        [6]   // Conveyor 6 Millisecond Accumulator Updated by STI File 18
        [7]   // Conveyor 7 Millisecond Accumulator Updated by STI File 18
        [8]   // Conveyor 8 Millisecond Accumulator Updated by STI File 18
        [9]   // Conveyor 9 Millisecond Accumulator Updated by STI File 18
        [16]   // Conveyor 16 Millisecond Accumulator Updated by STI File 18
        [17]   // Conveyor 17 Millisecond Accumulator Updated by STI File 18
        [18]   // Conveyor 18 Millisecond Accumulator Updated by STI File 18
        [19]   // Conveyor 19 Millisecond Accumulator Updated by STI File 18
        [20]   // conveyor 20 Millisecond Accumulator Updated by STI File 18
        [21]   // conveyor 21 Millisecond Accumulator Updated by STI File 18
        [22]   // conveyor 22 Millisecond Accumulator Updated by STI File 18
        [23]   // conveyor 23 Millisecond Accumulator Updated by STI File 18
        [24]   // conveyor 24 Millisecond Accumulator Updated by STI File 18
        [25]   // conveyor 25 Millisecond Accumulator Updated by STI File 18
        [26]   // conveyor 26 Millisecond Accumulator Updated by STI File 18
        [27]   // conveyor 27 Millisecond Accumulator Updated by STI File 18
        [28]   // conveyor 28 Millisecond Accumulator Updated by STI File 18
        [29]   // conveyor 29 Millisecond Accumulator Updated by STI File 18
        [30]   // conveyor 30 Millisecond Accumulator Updated by STI File 18
        [31]   // conveyor 31 Millisecond Accumulator Updated by STI File 18
   N301 : DINT[1];
   N302 : DINT[1];
   N303 : DINT[1];
   N304 : DINT[1];
   N305 : DINT[1];
   N306 : DINT[1];
   N307 : DINT[1];
   N308 : DINT[1];
   N309 : DINT[1];
   N31 : DINT[33];   // M2 to M4
        [1]   // Conveyor 1 Copy Buffer Transfers PLC IDs to Next Conveyor
        [2]   // Conveyor 2 Copy Buffer Transfers PLC IDs to Next Conveyor
        [3]   // Conveyor 3 Copy Buffer Transfers PLC IDs to Next Conveyor
        [4]   // Conveyor 4 Copy Buffer Transfers PLC IDs to Next Conveyor
        [5]   // Conveyor 5 Copy Buffer Transfers PLC IDs to Next Conveyor
        [6]   // Conveyor 6 Copy Buffer Transfers PLC IDs to Next Conveyor
        [7]   // Conveyor 7 Copy Buffer Transfers PLC IDs to Next Conveyor
        [8]   // Conveyor 8 Copy Buffer Transfers PLC IDs to Next Conveyor
        [9]   // Conveyor 9 Copy Buffer Transfers PLC IDs to Next Conveyor
        [10]   // Conveyor 10 Copy Buffer Transfers PLC IDs to Next Conveyor
        [11]   // Conveyor 11 Copy Buffer Transfers PLC IDs to Next Conveyor
        [12]   // Conveyor 12 Copy Buffer Transfers PLC IDs to Next Conveyor
        [13]   // Conveyor 13 Copy Buffer Transfers PLC IDs to Next Conveyor
        [14]   // Conveyor 14 Copy Buffer Transfers PLC IDs to Next Conveyor
        [15]   // Conveyor 15 Copy Buffer Transfers PLC IDs to Next Conveyor
        [16]   // Conveyor 16 Copy Buffer Transfers PLC IDs to Next Conveyor
        [17]   // Conveyor 17 Copy Buffer Transfers PLC IDs to Next Conveyor
        [18]   // Conveyor 18 Copy Buffer Transfers PLC IDs to Next Conveyor
        [19]   // Conveyor 19 Copy Buffer Transfers PLC IDs to Next Conveyor
        [20]   // Conveyor 20 Copy Buffer Transfers PLC IDs to Next Conveyor
        [21]   // Conveyor 21 Copy Buffer Transfers PLC IDs to Next Conveyor
        [22]   // Conveyor 22 Copy Buffer Transfers PLC IDs to Next Conveyor
        [23]   // Conveyor 23 Copy Buffer Transfers PLC IDs to Next Conveyor
        [24]   // Conveyor 24 Copy Buffer Transfers PLC IDs to Next Conveyor
        [25]   // Conveyor 25 Copy Buffer Transfers PLC IDs to Next Conveyor
        [26]   // Conveyor 26 Copy Buffer Transfers PLC IDs to Next Conveyor
        [27]   // Conveyor 27 Copy Buffer Transfers PLC IDs to Next Conveyor
        [28]   // Conveyor 28 Copy Buffer Transfers PLC IDs to Next Conveyor
        [29]   // Conveyor 29 Copy Buffer Transfers PLC IDs to Next Conveyor
        [30]   // Conveyor 30 Copy Buffer Transfers PLC IDs to Next Conveyor
        [31]   // Conveyor 31 Copy Buffer Transfers PLC IDs to Next Conveyor
        [32]   // Conveyor 32 Copy Buffer Transfers PLC IDs to Next Conveyor
   N310 : DINT[1];
   N311 : DINT[1];
   N312 : DINT[1];
   N313 : DINT[1];
   N314 : DINT[1];
   N315 : DINT[1];
   N316 : DINT[1];
   N317 : DINT[1];
   N318 : DINT[1];
   N319 : DINT[1];
   N32 : DINT[33] := ([0] := 1800, [1] := 67);
        [10]   // Conveyor 10 Tracking Zone Length
        [11]   // Conveyor 11 Tracking Zone Length
        [12]   // Conveyor 12 Tracking Zone Length
        [13]   // Conveyor 13 Tracking Zone Length
        [1]   // Conveyor 1 Tracking Zone Length
        [14]   // Conveyor 14 Tracking Zone Length
        [2]   // Conveyor 2 Tracking Zone Length
        [15]   // Conveyor 15 Tracking Zone Length
        [3]   // Conveyor 3 Tracking Zone Length
        [16]   // Conveyor 16 Tracking Zone Length
        [17]   // Conveyor 17 Tracking Zone Length
        [18]   // Conveyor 18 Tracking Zone Length
        [19]   // Conveyor 19 Tracking Zone Length
        [20]   // Conveyor 20 Tracking Zone Length
        [21]   // Conveyor 21 Tracking Zone Length
        [22]   // Conveyor 22 Tracking Zone Length
        [23]   // Conveyor 23 Tracking Zone Length
        [24]   // Conveyor 24 Tracking Zone Length
        [25]   // Conveyor 25 Tracking Zone Length
        [26]   // Conveyor 26 Tracking Zone Length
        [4]   // Conveyor 4 Tracking Zone Length
        [27]   // Conveyor 27 Tracking Zone Length
        [28]   // Conveyor 28 Tracking Zone Length
        [29]   // Conveyor 29 Tracking Zone Length
        [30]   // Conveyor 30 Tracking Zone Length
        [31]   // Conveyor 31 Tracking Zone Length
        [32]   // Conveyor 32 Tracking Zone Length
        [5]   // Conveyor 5 Tracking Zone Length
        [6]   // Conveyor 6 Tracking Zone Length
        [7]   // Conveyor 7 Tracking Zone Length
        [8]   // Conveyor 8 Tracking Zone Length
        [9]   // Conveyor 9 Tracking Zone Length
   N320 : DINT[1];
   N321 : DINT[1];
   N322 : DINT[1];
   N323 : DINT[1];
   N324 : DINT[1];
   N325 : DINT[1];
   N326 : DINT[1];
   N327 : DINT[1];
   N328 : DINT[1];
   N329 : DINT[1];
   N33 : DINT[2] := ([0] := 3000, [1] := 40);
   N330 : DINT[1];
   N331 : DINT[1];
   N332 : DINT[1];
   N334 : DINT[1];
   N335 : DINT[1];
   N336 : DINT[1];
   N337 : DINT[1];
   N338 : DINT[1];
   N339 : DINT[1];
   N340 : DINT[1];
   N341 : DINT[1];
   N342 : DINT[1];
   N343 : DINT[1];
   N344 : DINT[1];
   N345 : DINT[1];
   N346 : DINT[1];
   N347 : DINT[1];
   N348 : DINT[1];
   N349 : DINT[1];
   N35 : DINT[5] := ([0] := 32, [1] := 232, [2] := 33, [3] := 132, [4] := 24);
   N350 : DINT[1];
   N351 : DINT[1];
   N352 : DINT[1];
   N353 : DINT[1];
   N354 : DINT[1];
   N355 : DINT[1];
   N356 : DINT[1];
   N357 : DINT[1];
   N358 : DINT[1];
   N359 : DINT[1];
   N35_0 : ALIAS FOR N35[0];
   N35_1 : ALIAS FOR N35[1];
   N35_2 : ALIAS FOR N35[2];
   N35_4 : ALIAS FOR N35[4];
   N360 : DINT[1];
   N361 : DINT[1];
   N362 : DINT[1];
   N363 : DINT[1];
   N364 : DINT[1];
   N365 : DINT[1];
   N367 : DINT[1];
   N368 : DINT[1];
   N369 : DINT[1];
   N370 : DINT[1];
   N371 : DINT[1];
   N372 : DINT[1];
   N373 : DINT[1];
   N374 : DINT[1];
   N375 : DINT[1];
   N376 : DINT[1];
   N377 : DINT[1];
   N378 : DINT[1];
   N379 : DINT[1];
   N380 : DINT[1];
   N381 : DINT[1];
   N382 : DINT[1];
   N383 : DINT[1];
   N384 : DINT[1];
   N385 : DINT[1];
   N386 : DINT[1];
   N387 : DINT[1];
   N388 : DINT[1];
   N389 : DINT[1];
   N390 : DINT[1];
   N391 : DINT[1];
   N392 : DINT[1];
   N393 : DINT[1];
   N394 : DINT[1];
   N395 : DINT[1];
   N396 : DINT[1];
   N397 : DINT[1];
   N398 : DINT[1];
   N40 : DINT[32];
        [10]   // Conveyor 10 PLD ID of Cap being Resynced
        [11]   // Conveyor 11 PLD ID of Cap being Resynced
        [12]   // Conveyor 12 PLD ID of Cap being Resynced
        [13]   // Conveyor 13 PLD ID of Cap being Resynced
        [14]   // Conveyor 14 PLD ID of Cap being Resynced
        [15]   // Conveyor 15 PLD ID of Cap being Resynced
        [16]   // Conveyor 16 PLD ID of Cap being Resynced
        [17]   // Conveyor 17 PLD ID of Cap being Resynced
        [18]   // Conveyor 18 PLD ID of Cap being Resynced
        [19]   // Conveyor 19 PLD ID of Cap being Resynced
        [20]   // Conveyor 20 PLD ID of Cap being Resynced
        [21]   // Conveyor 21 PLD ID of Cap being Resynced
        [22]   // Conveyor 22 PLD ID of Cap being Resynced
        [23]   // Conveyor 23 PLD ID of Cap being Resynced
        [24]   // Conveyor 24 PLD ID of Cap being Resynced
        [25]   // Conveyor 25 PLD ID of Cap being Resynced
        [26]   // Conveyor 26 PLD ID of Cap being Resynced
        [27]   // Conveyor 27 PLD ID of Cap being Resynced
        [28]   // Conveyor 28 PLD ID of Cap being Resynced
        [29]   // Conveyor 29 PLD ID of Cap being Resynced
        [1]   // Conveyor 1 PLD ID of Cap being Resynced
        [2]   // Conveyor 2 PLD ID of Cap being Resynced
        [3]   // Conveyor 3 PLD ID of Cap being Resynced
        [4]   // Conveyor 4 PLD ID of Cap being Resynced
        [5]   // Conveyor 5 PLD ID of Cap being Resynced
        [6]   // Conveyor 6 PLD ID of Cap being Resynced
        [7]   // Conveyor 7 PLD ID of Cap being Resynced
        [8]   // Conveyor 8 PLD ID of Cap being Resynced
        [9]   // Conveyor 9 PLD ID of Cap being Resynced
        [30]   // Conveyor 30 PLD ID of Cap being Resynced
        [31]   // Conveyor 31 PLD ID of Cap being Resynced
   N400 : DINT[1];
   N401 : DINT[1];
   N402 : DINT[1];
   N403 : DINT[1];
   N404 : DINT[1];
   N405 : DINT[1];
   N406 : DINT[1];
   N407 : DINT[1];
   N408 : DINT[1];
   N409 : DINT[1];
   N410 : DINT[1];
   N411 : DINT[1];
   N412 : DINT[1];
   N413 : DINT[1];
   N414 : DINT[1];
   N415 : DINT[1];
   N416 : DINT[1];
   N417 : DINT[1];
   N418 : DINT[1];
   N419 : DINT[1];
   N420 : DINT[1];
   N421 : DINT[1];
   N422 : DINT[1];
   N423 : DINT[1];
   N424 : DINT[1];
   N425 : DINT[1];
   N426 : DINT[1];
   N427 : DINT[1];
   N428 : DINT[1];
   N429 : DINT[1];
   N430 : DINT[1];
   N431 : DINT[1];
   N433 : DINT[1];
   N434 : DINT[1];
   N435 : DINT[1];
   N436 : DINT[1];
   N437 : DINT[1];
   N438 : DINT[1];
   N439 : DINT[1];
   N440 : DINT[1];
   N441 : DINT[1];
   N442 : DINT[1];
   N443 : DINT[1];
   N444 : DINT[1];
   N445 : DINT[1];
   N446 : DINT[1];
   N447 : DINT[1];
   N448 : DINT[1];
   N449 : DINT[1];
   N450 : DINT[1];
   N451 : DINT[1];
   N452 : DINT[1];
   N453 : DINT[1];
   N454 : DINT[1];
   N455 : DINT[1];
   N456 : DINT[1];
   N457 : DINT[1];
   N458 : DINT[1];
   N459 : DINT[1];
   N460 : DINT[1];
   N461 : DINT[1];
   N462 : DINT[1];
   N463 : DINT[1];
   N464 : DINT[1];
   N466 : DINT[1];
   N467 : DINT[1];
   N468 : DINT[1];
   N469 : DINT[1];
   N470 : DINT[1];
   N471 : DINT[1];
   N472 : DINT[1];
   N473 : DINT[1];
   N474 : DINT[1];
   N475 : DINT[1];
   N476 : DINT[1];
   N477 : DINT[1];
   N478 : DINT[1];
   N479 : DINT[1];
   N480 : DINT[1];
   N481 : DINT[1];
   N482 : DINT[1];
   N483 : DINT[1];
   N484 : DINT[1];
   N485 : DINT[1];
   N486 : DINT[1];
   N487 : DINT[1];
   N488 : DINT[1];
   N489 : DINT[1];
   N490 : DINT[1];
   N491 : DINT[1];
   N492 : DINT[1];
   N493 : DINT[1];
   N494 : DINT[1];
   N495 : DINT[1];
   N496 : DINT[1];
   N497 : DINT[1];
   N500 : DINT[13] := ([1] := 1755, [2] := 1755, [3] := 1750, [4] := 1750, [5] := 1750, [6] := 1750, [7] := 1750, [8] := 1755, [9] := 1755, [10] := 1755, [11] := 1755, [12] := 1755);   // Motor RPM
        [10]   // M2CM10 Motor RPM
        [11]   // M2CM11 Motor RPM
        [12]   // M2CM12 Motor RPM
        [1]   // M2CM01 Motor RPM
        [2]   // M2CM02 Motor RPM
        [3]   // M2CM03 Motor RPM
        [4]   // M2CM04 Motor RPM
        [5]   // M2CM05 Motor RPM
        [6]   // M2CM06 Motor RPM
        [7]   // M2CM07 Motor RPM
        [8]   // M2CM08 Motor RPM
        [9]   // M2CM09 Motor RPM
   N501 : DINT[13] := ([1] := 43, [2] := 43, [3] := 43, [4] := 29, [5] := 29, [6] := 29, [7] := 29, [8] := 29, [9] := 29, [10] := 29, [11] := 29, [12] := 29);   // Gearbox raito
        [10]   // M2CM10 Gearbox raito
        [11]   // M2CM11 Gearbox raito
        [12]   // M2CM12 Gearbox raito
        [1]   // M2CM01 Gearbox raito
        [2]   // M2CM02 Gearbox raito
        [3]   // M2CM03 Gearbox raito
        [4]   // M2CM04 Gearbox raito
        [5]   // M2CM05 Gearbox raito
        [6]   // M2CM06 Gearbox raito
        [7]   // M2CM07 Gearbox raito
        [8]   // M2CM08 Gearbox raito
        [9]   // M2CM09 Gearbox raito
   N502 : DINT[13] := ([1] := 100, [2] := 100, [3] := 100, [4] := 100, [5] := 100, [6] := 100, [7] := 100, [8] := 100, [9] := 100, [10] := 100, [11] := 100, [12] := 100);   // Slip compensation
        [10]   // M2 CM10 Slip Compensation
        [11]   // M2 CM11 Slip Compensation
        [12]   // M2 CM12 Slip Compensation
        [1]   // M2 CM01 Slip Compensation
        [2]   // M2 CM02 Slip Compensation
        [3]   // M2 CM03 Slip Compensation
        [4]   // M2 CM04 Slip Compensation
        [5]   // M2 CM05 Slip Compensation
        [6]   // M2 CM06 Slip Compensation
        [7]   // M2 CM07 Slip Compensation
        [8]   // M2 CM08 Slip Compensation
        [9]   // M2 CM09 Slip Compensation
   N504 : DINT[13] := ([1] := 2042, [2] := 2042, [3] := 1728, [4] := 1728, [5] := 1728, [6] := 1728, [7] := 1728, [8] := 1728, [9] := 1728, [10] := 1728, [11] := 1728, [12] := 1728);   // Roll Circ
        [10]   // M2CM10 Roll Circ
        [11]   // M2CM11 Roll Circ
        [12]   // M2CM12 Roll Circ
        [1]   // M2CM01 Roll Circ
        [2]   // M2CM02 Roll Circ
        [3]   // M2CM03 Roll Circ
        [4]   // M2CM04 Roll Circ
        [5]   // M2CM05 Roll Circ
        [6]   // M2CM06 Roll Circ
        [7]   // M2CM07 Roll Circ
        [8]   // M2CM08 Roll Circ
        [9]   // M2CM09 Roll Circ
   N505 : DINT[13] := ([1] := 1397, [2] := 1397, [3] := 1179, [4] := 1748, [5] := 1748, [6] := 1748, [7] := 1748, [8] := 1753, [9] := 1753, [10] := 1753, [11] := 1753, [12] := 1753);   // IPM/HZ Conv Factor
        [10]   // M2CM10 IPM/HZ Conv Factor
        [11]   // M2CM11 IPM/HZ Conv Factor
        [12]   // M2CM12 IPM/HZ Conv Factor
        [1]   // M2CM01 IPM/HZ Conv Factor
        [2]   // M2CM02 IPM/HZ Conv Factor
        [3]   // M2CM03 IPM/HZ Conv Factor
        [4]   // M2CM04 IPM/HZ Conv Factor
        [5]   // M2CM05 IPM/HZ Conv Factor
        [6]   // M2CM06 IPM/HZ Conv Factor
        [7]   // M2CM07 IPM/HZ Conv Factor
        [8]   // M2CM08 IPM/HZ Conv Factor
        [9]   // M2CM09 IPM/HZ Conv Factor
   N507 : DINT[26] := ([1] := 94, [2] := 94, [3] := 112, [4] := 76, [5] := 76, [6] := 76, [7] := 76, [8] := 75, [9] := 75, [10] := 75, [11] := 75, [12] := 75, [13] := 322, [14] := 322, [15] := 382, [16] := 257, [17] := 257, [18] := 257, [19] := 257, [20] := 257, [21] := 257, [22] := 257, [23] := 257, [24] := 257, [25] := 450);   // Drive Command HZ
        [7]   // M2CM07S A1 Data In
   N54 : DINT[251];
   N601 : DINT[25];
   N602 : DINT[25];
   N603 : DINT[25];
   N604 : DINT[25];
   N605 : DINT[25];
   N606 : DINT[25];
   N607 : DINT[25];
   N608 : DINT[25];
   N609 : DINT[25];
   N610 : DINT[25];
   N611 : DINT[25];
   N612 : DINT[25];
   N613 : DINT[25];
   N614 : DINT[25];
   N615 : DINT[25];
   N616 : DINT[25];
   N617 : DINT[25];
   N618 : DINT[25];
   N619 : DINT[25];
   N620 : DINT[25];
   N621 : DINT[25];
   N622 : DINT[25];
   N623 : DINT[25];
   N624 : DINT[25];
   N625 : DINT[25];
   N626 : DINT[25];
   N627 : DINT[25];
   N628 : DINT[25];
   N629 : DINT[25];
   N630 : DINT[25];
   N631 : DINT[25];
   N632 : DINT[25];
   N633 : DINT[25];
   N634 : DINT[25];
   N635 : DINT[25];
   N636 : DINT[25];
   N637 : DINT[25];
   N638 : DINT[25];
   N639 : DINT[25];
   N640 : DINT[25];
   N641 : DINT[25];
   N642 : DINT[25];
   N643 : DINT[25];
   N644 : DINT[25];
   N645 : DINT[25];
   N646 : DINT[25];
   N647 : DINT[25];
   N648 : DINT[25];
   N649 : DINT[25];
   N650 : DINT[25];
   N651 : DINT[25];
   N652 : DINT[25];
   N653 : DINT[25];
   N654 : DINT[25];
   N655 : DINT[25];
   N656 : DINT[25];
   N657 : DINT[25];
   N658 : DINT[25];
   N659 : DINT[25];
   N660 : DINT[25];
   N662 : DINT[25];
   N663 : DINT[25];
   N664 : DINT[25];
   N665 : DINT[25];
   N666 : DINT[25];
   N667 : DINT[25];
   N668 : DINT[25];
   N669 : DINT[25];
   N670 : DINT[25];
   N671 : DINT[25];
   N672 : DINT[25];
   N673 : DINT[25];
   N674 : DINT[25];
   N675 : DINT[25];
   N676 : DINT[25];
   N677 : DINT[25];
   N678 : DINT[25];
   N679 : DINT[25];
   N680 : DINT[25];
   N681 : DINT[25];
   N682 : DINT[25];
   N683 : DINT[25];
   N684 : DINT[25];
   N685 : DINT[25];
   N686 : DINT[25];
   N687 : DINT[25];
   N688 : DINT[25];
   N689 : DINT[25];
   N690 : DINT[25];
   N691 : DINT[25];
   N692 : DINT[25];
   N693 : DINT[25];
   N694 : DINT[25];
   N695 : DINT[25];
   N696 : DINT[25];
   N697 : DINT[25];
   N698 : DINT[25];
   N699 : DINT[25];
   N7 : DINT[101] := ([10] := 3500, [11] := 100, [20] := 3930);
        [10]   // Current Command Frequency
        [0]   // DH+ Station number set on processor DIP switches
        [11]   // Current Test Addition Operand
   N70 : DINT[128] := ([0] := 11008);
   N700 : DINT[25];
   N701 : DINT[25];
   N702 : DINT[25];
   N703 : DINT[25];
   N704 : DINT[25];
   N705 : DINT[25];
   N706 : DINT[25];
   N707 : DINT[25];
   N708 : DINT[25];
   N709 : DINT[25];
   N71 : DINT[128] := ([2] := 40, [4] := 60);
        [2]   // M2CM12 A1 Data In
        [4]   // M2CM12 A2 Data In
   N710 : DINT[25];
   N711 : DINT[25];
   N712 : DINT[25];
   N713 : DINT[25];
   N714 : DINT[25];
   N715 : DINT[25];
   N716 : DINT[25];
   N717 : DINT[25];
   N718 : DINT[25];
   N719 : DINT[25];
   N72 : DINT[200] := ([0] := 4095);
        [0].0   // M2CM01 Drive Healthy and Running
        [0].1   // M2CM02 Drive Healthy and Running
        [0].2   // M2CM03 Drive Healthy and Running
        [3]   // VMCC M2 Drive Fault or Not Running Bits NORTH
        [0]   // VMCC M2 Drive Status Word Drive Healthy
        [1]   // VMCC M2 Drive Fault or Not Running Bits
        [0].10   // M2CM11 Drive Healthy and Running
        [0].11   // M2CM12 Drive Healthy and Running
        [2].10   // M2CM11N Drive Healthy and Running
        [2].11   // M2CM12N Drive Healthy and Running
        [0].3   // M2CM04 Drive Healthy and Running
        [0].4   // M2CM05 Drive Healthy and Running
        [0].5   // M2CM06 Drive Healthy and Running
        [0].6   // M2CM07 Drive Healthy and Running
        [0].7   // M2CM08 Drive Healthy and Running
        [0].8   // M2CM09 Drive Healthy and Running
        [0].9   // M2CM10 Drive Healthy and Running
        [2].3   // M2CM04N Drive Healthy and Running
        [2].4   // M2CM05N Drive Healthy and Running
        [2].5   // M2CM06N Drive Healthy and Running
        [2].6   // M2CM07N Drive Healthy and Running
        [2].7   // M2CM08N Drive Healthy and Running
        [2].8   // M2CM09N Drive Healthy and Running
        [2].9   // M2CM10N Drive Healthy and Running
   N720 : DINT[25];
   N721 : DINT[25];
   N723 : DINT[25];
   N724 : DINT[25];
   N725 : DINT[25];
   N726 : DINT[25];
   N727 : DINT[25];
   N728 : DINT[25];
   N729 : DINT[25];
   N730 : DINT[25];
   N731 : DINT[25];
   N732 : DINT[25];
   N733 : DINT[25];
   N734 : DINT[25];
   N735 : DINT[25];
   N736 : DINT[25];
   N737 : DINT[25];
   N738 : DINT[25];
   N739 : DINT[25];
   N740 : DINT[25];
   N741 : DINT[25];
   N742 : DINT[25];
   N743 : DINT[25];
   N744 : DINT[25];
   N745 : DINT[25];
   N746 : DINT[25];
   N747 : DINT[25];
   N748 : DINT[25];
   N749 : DINT[25];
   N750 : DINT[25];
   N751 : DINT[25];
   N752 : DINT[25];
   N753 : DINT[25];
   N754 : DINT[25];
   N755 : DINT[25];
   N756 : DINT[25];
   N758 : DINT[25];
   N759 : DINT[25];
   N760 : DINT[25];
   N761 : DINT[25];
   N762 : DINT[25];
   N763 : DINT[25];
   N764 : DINT[25];
   N765 : DINT[25];
   N766 : DINT[25];
   N767 : DINT[25];
   N768 : DINT[25];
   N769 : DINT[25];
   N770 : DINT[25];
   N771 : DINT[25];
   N772 : DINT[25];
   N773 : DINT[25];
   N774 : DINT[25];
   N775 : DINT[25];
   N776 : DINT[25];
   N777 : DINT[25];
   N778 : DINT[25];
   N779 : DINT[25];
   N780 : DINT[25];
   N781 : DINT[25];
   N782 : DINT[25];
   N783 : DINT[25];
   N784 : DINT[25];
   N785 : DINT[25];
   N786 : DINT[25];
   N787 : DINT[25];
   N788 : DINT[25];
   N789 : DINT[25];
   N790 : DINT[25];
   N791 : DINT[25];
   N792 : DINT[25];
   N793 : DINT[25];
   N794 : DINT[25];
   N795 : DINT[25];
   N796 : DINT[25];
   N797 : DINT[25];
   N798 : DINT[25];
   N799 : DINT[25];
   N80 : DINT[65] := ([11] := 2415, [12] := 5642, [15] := 2284, [16] := 5646, [19] := 1825, [20] := 4512, [23] := 1683, [24] := 4510, [27] := 1685, [28] := 4515, [31] := 1682, [32] := 4517, [35] := 1697, [36] := 452, [39] := 1681, [40] := 2811, [43] := 1681, [44] := 2811, [47] := 1681, [48] := 2811, [51] := 1684, [52] := 2815, [55] := 3995, [56] := 5974, [60] := 3000, [64] := 3000);
        [13].8   // M2CM02 Accel Time
        [1]   // RIO SN WRITE DATA Reserved Not Used
        [13].9   // M2CM02 Accel Time
        [2]   // RIO SN WRITE DATA Reserved Not Used
        [13].1   // M2CM02 Start
        [13]   // M2CM02 Drive Command
        [3]   // RIO SN WRITE DATA Reserved Not Used
        [4]   // RIO SN WRITE DATA Reserved Not Used
        [13].6   // M2CM02 Local
        [17].1   // M2CM03 Start
        [9].8   // M2CM01 Accel Time
        [9].9   // M2CM01 Accel Time
        [13].7   // M2CM02 MOP Increment
        [10]   // M2CM01 Speed Reference
        [5]   // RIO SN WRITE DATA Reserved Not Used
        [6]   // RIO SN WRITE DATA Reserved Not Used
        [7]   // RIO SN WRITE DATA Reserved Not Used
        [13].15   // M2CM02 MOP Decrement
        [8]   // RIO SN WRITE DATA Reserved Not Used
        [17].8   // M2CM03 Accel Time
        [17].15   // M2CM03 MOP Decrement
        [21].15   // M2CM04 MOP Decrement
        [25].15   // M2CM05 MOP Decrement
        [18].1   // M2CM03 Reference Select
        [13].12   // M2CM02 Reference Select
        [13].13   // M2CM02 Reference Select
        [13].14   // M2CM02 Reference Select
        [13].0   // M2CM02 Stop
        [17].0   // M2CM03 Stop
        [14]   // M2CM02 Speed Reference
        [11]   // M2CM01 A1 Data In
        [12]   // M2CM01 A2 Data In
        [13].4   // M2CM02 Direction
        [21].0   // M2CM04 Stop
        [17].6   // M2CM03 Local
        [13].10   // M2CM02 Decel Time
        [13].11   // M2CM02 Decel Time
        [17].12   // M2CM03 Reference Select
        [17].13   // M2CM03 Reference Select
        [17].14   // M2CM03 Reference Select
        [29].15   // M2CM06 MOP Decrement
        [13].2   // M2CM02 Jog
        [13].3   // M2CM02 Clear Faults
        [13].5   // M2CM02 Direction
        [17]   // M2CM03 Drive Command
        [21].1   // M2CM04 Start
        [17].7   // M2CM03 MOP Increment
        [17].9   // M2CM03 Accel Time
        [21].8   // M2CM04 Accel Time
        [18]   // M2CM03 Speed Reference
        [15]   // M2CM02 A1 Data In
        [16]   // M2CM02 A2 Data In
        [17].4   // M2CM03 Direction
        [25].0   // M2CM05 Stop
        [21].6   // M2CM04 Local
        [17].10   // M2CM03 Decel Time
        [17].11   // M2CM03 Decel Time
        [21].12   // M2CM04 Reference Select
        [21].13   // M2CM04 Reference Select
        [21].14   // M2CM04 Reference Select
        [33].15   // M2CM07 MOP Decrement
        [17].2   // M2CM03 Jog
        [17].3   // M2CM03 Clear Faults
        [17].5   // M2CM03 Direction
        [21]   // M2CM04 Drive Command
        [25].1   // M2CM05 Start
        [21].7   // M2CM04 MOP Increment
        [21].9   // M2CM04 Accel Time
        [25].8   // M2CM05 Accel Time
        [22]   // M2CM04 Speed Reference
        [22].5   // M2CM04 Reference Select
        [19]   // M2CM03 A1 Data In
        [20]   // M2CM03 A2 Data In
        [21].4   // M2CM04 Direction
        [29].0   // M2CM06 Stop
        [25].6   // M2CM05 Local
        [21].10   // M2CM04 Decel Time
        [21].11   // M2CM04 Decel Time
        [25].12   // M2CM05 Reference Select
        [25].13   // M2CM05 Reference Select
        [25].14   // M2CM05 Reference Select
        [37].15   // M2CM08 MOP Decrement
        [21].2   // M2CM04 Jog
        [21].3   // M2CM04 Clear Faults
        [21].5   // M2CM04 Direction
        [25]   // M2CM05 Drive Command
        [29].1   // M2CM06 Start
        [25].7   // M2CM05 MOP Increment
        [25].9   // M2CM05 Accel Time
        [29].8   // M2CM06 Accel Time
        [26]   // M2CM05 Speed Reference
        [26].9   // M2CM05 Reference Select
        [23]   // M2CM04 A1 Data In
        [24]   // M2CM04 A2 Data In
        [25].4   // M2CM05 Direction
        [33].0   // M2CM07 Stop
        [29].6   // M2CM06 Local
        [25].10   // M2CM05 Decel Time
        [25].11   // M2CM05 Decel Time
        [29].12   // M2CM06 Reference Select
        [29].13   // M2CM06 Reference Select
        [29].14   // M2CM06 Reference Select
        [41].15   // M2CM09 MOP Decrement
        [25].2   // M2CM05 Jog
        [25].3   // M2CM05 Clear Faults
        [25].5   // M2CM05 Direction
        [29]   // M2CM06 Drive Command
        [33].1   // M2CM07 Start
        [29].7   // M2CM06 MOP Increment
        [29].9   // M2CM06 Accel Time
        [33].8   // M2CM07 Accel Time
        [30]   // M2CM06 Speed Reference
        [35].1   // M2CM07 Reference Select
        [27]   // M2CM05 A1 Data In
        [28]   // M2CM05 A2 Data In
        [29].4   // M2CM06 Direction
        [37].0   // M2CM08 Stop
        [33].6   // M2CM07 Local
        [29].10   // M2CM06 Decel Time
        [29].11   // M2CM06 Decel Time
        [30].13   // M2CM06 Reference Select
        [33].12   // M2CM07 Reference Select
        [33].13   // M2CM07 Reference Select
        [45].15   // M2CM10 MOP Decrement
        [29].2   // M2CM06 Jog
        [29].3   // M2CM06 Clear Faults
        [29].5   // M2CM06 Direction
        [33]   // M2CM07 Drive Command
        [37].1   // M2CM08 Start
        [33].7   // M2CM07 MOP Increment
        [33].9   // M2CM07 Accel Time
        [37].8   // M2CM08 Accel Time
        [34]   // M2CM07 Speed Reference
        [33].14   // M2CM07 Reference Select
        [31]   // M2CM06 A1 Data In
        [32]   // M2CM06 A2 Data In
        [33].4   // M2CM07 Direction
        [41].0   // M2CM09 Stop
        [37].6   // M2CM08 Local
        [33].10   // M2CM07 Decel Time
        [33].11   // M2CM07 Decel Time
        [37].12   // M2CM08 Reference Select
        [37].13   // M2CM08 Reference Select
        [37].14   // M2CM08 Reference Select
        [49].15   // M2CM11 MOP Decrement
        [33].2   // M2CM07 Jog
        [33].3   // M2CM07 Clear Faults
        [33].5   // M2CM07 Direction
        [37]   // M2CM08 Drive Command
        [41].1   // M2CM09 Start
        [37].7   // M2CM08 MOP Increment
        [37].9   // M2CM08 Accel Time
        [41].8   // M2CM09 Accel Time
        [38]   // M2CM08 Speed Reference
        [35]   // M2CM07 A1 Data In
        [39].5   // M2CM08 Reference Select
        [36]   // M2CM07 A2 Data In
        [37].4   // M2CM08 Direction
        [45].0   // M2CM10 Stop
        [41].6   // M2CM09 Local
        [37].10   // M2CM08 Decel Time
        [37].11   // M2CM08 Decel Time
        [41].12   // M2CM09 Reference Select
        [41].13   // M2CM09 Reference Select
        [41].14   // M2CM09 Reference Select
        [53].15   // M2CM12 MOP Decrement
        [37].2   // M2CM08 Jog
        [37].3   // M2CM08 Clear Faults
        [37].5   // M2CM08 Direction
        [41]   // M2CM09 Drive Command
        [45].1   // M2CM10 Start
        [41].7   // M2CM09 MOP Increment
        [41].9   // M2CM09 Accel Time
        [45].8   // M2CM10 Accel Time
        [42]   // M2CM09 Speed Reference
        [39]   // M2CM08 A1 Data In
        [43].9   // M2CM09 Reference Select
        [40]   // M2CM08 A2 Data In
        [41].4   // M2CM09 Direction
        [49].0   // M2CM11 Stop
        [45].6   // M2CM10 Local
        [41].10   // M2CM09 Decel Time
        [41].11   // M2CM09 Decel Time
        [45].12   // M2CM10 Reference Select
        [45].13   // M2CM10 Reference Select
        [45].14   // M2CM10 Reference Select
        [41].2   // M2CM09 Jog
        [41].3   // M2CM09 Clear Faults
        [41].5   // M2CM09 Direction
        [45]   // M2CM10 Drive Command
        [49].1   // M2CM11 Start
        [45].7   // M2CM10 MOP Increment
        [45].9   // M2CM10 Accel Time
        [49].8   // M2CM11 Accel Time
        [46]   // M2CM10 Speed Reference
        [43]   // M2CM09 A1 Data In
        [52].1   // M2CM11 Reference Select
        [44]   // M2CM09 A2 Data In
        [45].4   // M2CM10 Direction
        [53].0   // M2CM12 Stop
        [49].6   // M2CM11 Local
        [45].10   // M2CM10 Decel Time
        [45].11   // M2CM10 Decel Time
        [47].13   // M2CM10 Reference Select
        [49].12   // M2CM11 Reference Select
        [49].13   // M2CM11 Reference Select
        [45].2   // M2CM10 Jog
        [45].3   // M2CM10 Clear Faults
        [45].5   // M2CM10 Direction
        [49]   // M2CM11 Drive Command
        [53].1   // M2CM12 Start
        [49].7   // M2CM11 MOP Increment
        [49].9   // M2CM11 Accel Time
        [53].8   // M2CM12 Accel Time
        [50]   // M2CM11 Speed Reference
        [47]   // M2CM10 A1 Data In
        [49].14   // M2CM11 Reference Select
        [48]   // M2CM10 A2 Data In
        [49].4   // M2CM11 Direction
        [53].6   // M2CM12 Local
        [49].10   // M2CM11 Decel Time
        [49].11   // M2CM11 Decel Time
        [53].12   // M2CM12 Reference Select
        [53].13   // M2CM12 Reference Select
        [53].14   // M2CM12 Reference Select
        [49].2   // M2CM11 Jog
        [49].3   // M2CM11 Clear Faults
        [49].5   // M2CM11 Direction
        [53]   // M2CM12 Drive Command
        [53].7   // M2CM12 MOP Increment
        [53].9   // M2CM12 Accel Time
        [9].10   // M2CM01 Decel Time
        [54]   // M2CM12 Speed Reference
        [51]   // M2CM11 A1 Data In
        [52]   // M2CM11 A2 Data In
        [56].5   // M2CM12 Reference Select
        [53].4   // M2CM12 Direction
        [53].10   // M2CM12 Decel Time
        [53].11   // M2CM12 Decel Time
        [53].2   // M2CM12 Jog
        [53].3   // M2CM12 Clear Faults
        [53].5   // M2CM12 Direction
        [9].15   // M2CM01 MOP Decrement
        [9].11   // M2CM01 Decel Time
        [9].3   // M2CM01 Clear Faults
        [9].7   // M2CM01 MOP Increment
        [55]   // M2CM12 A1 Data In
        [56]   // M2CM12 A2 Data In
        [9].12   // M2CM01 Reference Select
        [9]   // M2CM01 Drive Command
        [9].0   // M2CM01 Stop
        [9].1   // M2CM01 Start
        [9].13   // M2CM01 Reference Select
        [9].14   // M2CM01 Reference Select
        [9].2   // M2CM01 Jog
        [9].4   // M2CM01 Direction
        [9].5   // M2CM01 Direction
        [9].6   // M2CM01 Local
   N802 : INT[420] := ([2] := 95, [4] := 322, [22] := 95, [24] := 322, [42] := 113, [44] := 382, [62] := 76, [64] := 256, [82] := 76, [84] := 257, [102] := 76, [104] := 256, [122] := 76, [124] := 257, [142] := 76, [144] := 256, [162] := 76, [164] := 257, [182] := 76, [184] := 256, [202] := 72, [204] := 243, [222] := 76, [224] := 256, [242] := 76, [244] := 257, [262] := 76, [264] := 256, [282] := 76, [284] := 257, [302] := 76, [304] := 257, [322] := 76, [324] := 257, [342] := 76, [344] := 258, [362] := 76, [364] := 257, [382] := 76, [384] := 258, [402] := 76, [404] := 257);
        [202]   // M2CM07N A1 Data In Changed logic to control speed of CM07N;28Mar2019,AAC
        [204]   // M2CM7N A2 Data In Changed logic to control speed of CM07N;28Mar2019,AAC
        [2]   // M2CM01 A1 Data In
        [4]   // M2CM01 A2 Data In
        [104]   // M2CM5S A2 Data In
        [124]   // M2CM5N A2 Data In
        [144]   // M2CM6S A2 Data In
        [102]   // M2CM05S A1 Data In
        [122]   // M2CM05N A1 Data In
        [164]   // M2CM6N A2 Data In
        [142]   // M2CM06S A1 Data In
        [184]   // M2CM7S A2 Data In
        [162]   // M2CM06N A1 Data In
        [224]   // M2CM8S A2 Data In
        [182]   // M2CM07S A1 Data In
        [244]   // M2CM8N A2 Data In
        [222]   // M2CM08S A1 Data In
        [262]   // M2CM9S A1 Data In
        [242]   // M2CM08N A1 Data In
        [264]   // M2CM9S A2 Data In
        [22]   // M2CM02 A1 Data In
        [302]   // M2CM10S A1 Data In
        [282]   // M2CM9N A1 Data In
        [24]   // M2CM02 A2 Data In
        [284]   // M2CM9N A2 Data In
        [304]   // M2CM10S A2 Data In
        [322]   // M2CM10N A1 Data In
        [324]   // M2CM10N A2 Data In
        [342]   // M2CM11S A1 Data In
        [344]   // M2CM11S A2 Data In
        [362]   // M2CM11N A1 Data In
        [364]   // M2CM11N A2 Data In
        [382]   // M2CM12S A1 Data In
        [384]   // M2CM12S A2 Data In
        [402]   // M2CM12N A1 Data In
        [404]   // M2CM12N A2 Data In
        [42]   // M2CM03 A1 Data In
        [44]   // M2CM03 A2 Data In
        [62]   // M2CM04S A1 Data In
        [64]   // M2CM4S A2 Data In
        [82]   // M2CM04N A1 Data In
        [84]   // M2CM4N A2 Data In
   N803 : INT[420] := ([0] := 2394, [2] := 4, [20] := 2394, [22] := 4, [40] := 2823, [42] := 4, [60] := 1915, [62] := 4, [80] := 1914, [82] := 4, [100] := 1915, [102] := 4, [120] := 1915, [122] := 4, [140] := 6452, [142] := 4, [160] := 6478, [162] := 4, [180] := 6452, [182] := 4, [200] := 6125, [202] := 4, [220] := 6452, [222] := 4, [240] := 6478, [242] := 4, [260] := 6452, [262] := 4, [280] := 6478, [282] := 4, [300] := 6478, [302] := 4, [320] := 6478, [322] := 4, [340] := 12124, [342] := 75, [360] := 12073, [362] := 75, [380] := 12124, [382] := 75, [400] := 12073, [402] := 75);
        [302]   // Check for 20 Comm-R Comms fault M2CM10S
        [2]   // Check for 20 Comm-R Comms fault M2CM01
        [322]   // Check for 20 Comm-R Comms fault M2CM10N
        [22]   // Check for 20 Comm-R Comms fault M2CM2
        [42]   // Check for 20 Comm-R Comms fault M2CM3
        [102]   // Check for 20 Comm-R Comms fault M2CM5S
        [342]   // Check for 20 Comm-R Comms fault M2CM11S
        [362]   // Check for 20 Comm-R Comms fault M2CM11N
        [382]   // Check for 20 Comm-R Comms fault M2CM12S
        [402]   // Check for 20 Comm-R Comms fault M2CM12N
        [122]   // Check for 20 Comm-R Comms fault M2CM5N
        [142]   // Check for 20 Comm-R Comms fault M2CM6S
        [162]   // Check for 20 Comm-R Comms fault M2CM6N
        [182]   // Check for 20 Comm-R Comms fault M2CM7S
        [202]   // Check for 20 Comm-R Comms fault M2CM7N
        [222]   // Check for 20 Comm-R Comms fault M2CM8S
        [242]   // Check for 20 Comm-R Comms fault M2CM8N
        [262]   // Check for 20 Comm-R Comms fault M2CM9S
        [282]   // Check for 20 Comm-R Comms fault M2CM9N
        [62]   // Check for 20 Comm-R Comms fault M2CM4S
        [82]   // Check for 20 Comm-R Comms fault M2CM4N
        [40]   // Block READ for M2CM2
   N81 : DINT[65] := ([6] := 14337, [7] := -1, [8] := -3841);
        [8].10   // RIO SN READ DATA Reserved Not Used
        [8].8   // RIO SN READ DATA Reserved Not Used
        [8].9   // RIO SN READ DATA Reserved Not Used
        [7].10   // RIO SN READ DATA Rack 4 Groups 2 and 3 Fault Bt
        [7].11   // RIO SN READ DATA Rack 4 Groups 0 and 1 Fault Bt
        [7].12   // RIO SN READ DATA Rack 3 Groups 6 and 7 Fault Bt
        [7].13   // RIO SN READ DATA Rack 3 Groups 4 and 5 Fault Bt
        [7].14   // RIO SN READ DATA Rack 3 Groups 2 and 3 Fault Bt
        [7].15   // RIO SN READ DATA Rack 3 Groups 0 and 1 Fault Bt
        [8].12   // RIO SN READ DATA Rack 7 Groups 6 and 7 Fault Bt
        [8].13   // RIO SN READ DATA Rack 7 Groups 4 and 5 Fault Bt
        [8].14   // RIO SN READ DATA Rack 7 Groups 2 and 3 Fault Bt
        [8].15   // RIO SN READ DATA Rack 7 Groups 0 and 1 Fault Bt
        [7].0   // RIO SN READ DATA Rack 2 Groups 6 and 7 Fault Bt
        [7].1   // RIO SN READ DATA Rack 2 Groups 4 and 5 Fault Bt
        [7].2   // RIO SN READ DATA Rack 2 Groups 2 and 3 Fault Bt
        [7].3   // RIO SN READ DATA Rack 2 Groups 0 and 1 Fault Bt
        [7].4   // RIO SN READ DATA Rack 1 Groups 6 and 7 Fault Bt
        [7].5   // RIO SN READ DATA Rack 1 Groups 4 and 5 Fault Bt
        [7].6   // RIO SN READ DATA Rack 1 Groups 2 and 3 Fault Bt
        [8].11   // RIO SN READ DATA Reserved Not Used
        [7].7   // RIO SN READ DATA Rack 1 Groups 0 and 1 Fault Bt
        [7].8   // RIO SN READ DATA Rack 4 Groups 6 and 7 Fault Bt
        [7].9   // RIO SN READ DATA Rack 4 Groups 4 and 5 Fault Bt
        [8].0   // RIO SN READ DATA Rack 6 Groups 6 and 7 Fault Bt
        [13]   // M2CM02 Drive Status
        [13].12   // M2CM02 Reference ID
        [8].1   // RIO SN READ DATA Rack 6 Groups 4 and 5 Fault Bt
        [8].2   // RIO SN READ DATA Rack 6 Groups 2 and 3 Fault Bt
        [8].3   // RIO SN READ DATA Rack 6 Groups 0 and 1 Fault Bt
        [8].4   // RIO SN READ DATA Rack 5 Groups 6 and 7 Fault Bt
        [8].5   // RIO SN READ DATA Rack 5 Groups 4 and 5 Fault Bt
        [8].6   // RIO SN READ DATA Rack 5 Groups 2 and 3 Fault Bt
        [8].7   // RIO SN READ DATA Rack 5 Groups 0 and 1 Fault Bt
        [1]   // RIO SN READ DATA Reserved Not Used
        [2]   // RIO SN READ DATA Reserved Not Used
        [3]   // RIO SN READ DATA Reserved Not Used
        [4]   // RIO SN READ DATA Reserved Not Used
        [5]   // RIO SN READ DATA Reserved Not Used
        [6]   // RIO SN READ DATA Reserved Fault Count
        [13].6   // M2CM02 Alarm
        [17].6   // M2CM03 Alarm
        [13].10   // M2CM02 Local Adaptor ID
        [13].11   // M2CM02 Local Adaptor ID
        [17].10   // M2CM03 Local Adaptor ID
        [21].6   // M2CM04 Alarm
        [9].4   // M2CM01 Accelerating
        [9].5   // M2CM01 Decelerating
        [13].3   // M2CM02 Actual Direction
        [13].2   // M2CM02 Cmd Direction
        [10]   // M2CM01 Speed Reference
        [13].8   // M2CM02 At Speed
        [17]   // M2CM03 Drive Status
        [14]   // M2CM02 Speed Reference
        [11]   // M2CM01 A1 Data Out
        [12]   // M2CM01 A2 Data Out
        [17].8   // M2CM03 At Speed
        [13].0   // M2CM02 Enabled
        [13].1   // M2CM02 Running
        [17].11   // M2CM03 Local Adaptor ID
        [21].10   // M2CM04 Local Adaptor ID
        [13].13   // M2CM02 Reference ID
        [13].14   // M2CM02 Reference ID
        [13].15   // M2CM02 Reference ID
        [17].12   // M2CM03 Reference ID
        [17].2   // M2CM03 Cmd Direction
        [13].9   // M2CM02 Local Adaptor ID
        [13].4   // M2CM02 Accelerating
        [13].5   // M2CM02 Decelerating
        [25].6   // M2CM05 Alarm
        [13].7   // M2CM02 Faulted
        [21]   // M2CM04 Drive Status
        [17].3   // M2CM03 Actual Direction
        [18]   // M2CM03 Speed Reference
        [15]   // M2CM02 A1 Data Out
        [16]   // M2CM02 A2 Data Out
        [21].8   // M2CM04 At Speed
        [17].0   // M2CM03 Enabled
        [17].1   // M2CM03 Running
        [21].11   // M2CM04 Local Adaptor ID
        [25].10   // M2CM05 Local Adaptor ID
        [17].13   // M2CM03 Reference ID
        [17].14   // M2CM03 Reference ID
        [17].15   // M2CM03 Reference ID
        [21].12   // M2CM04 Reference ID
        [21].2   // M2CM04 Cmd Direction
        [17].9   // M2CM03 Local Adaptor ID
        [17].4   // M2CM03 Accelerating
        [17].5   // M2CM03 Decelerating
        [29].6   // M2CM06 Alarm
        [17].7   // M2CM03 Faulted
        [25]   // M2CM05 Drive Status
        [21].3   // M2CM04 Actual Direction
        [22]   // M2CM04 Speed Reference
        [18].1   // M2CM03 Reference ID
        [19]   // M2CM03 A1 Data Out
        [20]   // M2CM03 A2 Data Out
        [25].8   // M2CM05 At Speed
        [21].0   // M2CM04 Enabled
        [21].1   // M2CM04 Running
        [25].11   // M2CM05 Local Adaptor ID
        [29].10   // M2CM06 Local Adaptor ID
        [21].13   // M2CM04 Reference ID
        [21].14   // M2CM04 Reference ID
        [21].15   // M2CM04 Reference ID
        [25].12   // M2CM05 Reference ID
        [25].2   // M2CM05 Cmd Direction
        [21].9   // M2CM04 Local Adaptor ID
        [21].4   // M2CM04 Accelerating
        [21].5   // M2CM04 Decelerating
        [33].6   // M2CM07 Alarm
        [21].7   // M2CM04 Faulted
        [29]   // M2CM06 Drive Status
        [25].3   // M2CM05 Actual Direction
        [26]   // M2CM05 Speed Reference
        [22].5   // M2CM04 Reference ID
        [23]   // M2CM04 A1 Data Out
        [24]   // M2CM04 A2 Data Out
        [29].8   // M2CM06 At Speed
        [25].0   // M2CM05 Enabled
        [25].1   // M2CM05 Running
        [29].11   // M2CM06 Local Adaptor ID
        [33].10   // M2CM07 Local Adaptor ID
        [25].13   // M2CM05 Reference ID
        [25].14   // M2CM05 Reference ID
        [25].15   // M2CM05 Reference ID
        [29].12   // M2CM06 Reference ID
        [29].2   // M2CM06 Cmd Direction
        [25].9   // M2CM05 Local Adaptor ID
        [25].4   // M2CM05 Accelerating
        [25].5   // M2CM05 Decelerating
        [37].6   // M2CM08 Alarm
        [25].7   // M2CM05 Faulted
        [33]   // M2CM07 Drive Status
        [29].3   // M2CM06 Actual Direction
        [30]   // M2CM06 Speed Reference
        [26].9   // M2CM05 Reference ID
        [27]   // M2CM05 A1 Data Out
        [28]   // M2CM05 A2 Data Out
        [33].8   // M2CM07 At Speed
        [29].0   // M2CM06 Enabled
        [29].1   // M2CM06 Running
        [33].11   // M2CM07 Local Adaptor ID
        [37].10   // M2CM08 Local Adaptor ID
        [29].13   // M2CM06 Reference ID
        [29].14   // M2CM06 Reference ID
        [29].15   // M2CM06 Reference ID
        [30].13   // M2CM06 Reference ID
        [33].2   // M2CM07 Cmd Direction
        [29].9   // M2CM06 Local Adaptor ID
        [29].4   // M2CM06 Accelerating
        [29].5   // M2CM06 Decelerating
        [41].6   // M2CM09 Alarm
        [29].7   // M2CM06 Faulted
        [37]   // M2CM08 Drive Status
        [33].3   // M2CM07 Actual Direction
        [34]   // M2CM07 Speed Reference
        [33].12   // M2CM07 Reference ID
        [31]   // M2CM06 A1 Data Out
        [32]   // M2CM06 A2 Data Out
        [37].8   // M2CM08 At Speed
        [33].0   // M2CM07 Enabled
        [33].1   // M2CM07 Running
        [37].11   // M2CM08 Local Adaptor ID
        [41].10   // M2CM09 Local Adaptor ID
        [33].13   // M2CM07 Reference ID
        [33].14   // M2CM07 Reference ID
        [33].15   // M2CM07 Reference ID
        [37].12   // M2CM08 Reference ID
        [37].2   // M2CM08 Cmd Direction
        [33].9   // M2CM07 Local Adaptor ID
        [33].4   // M2CM07 Accelerating
        [33].5   // M2CM07 Decelerating
        [45].6   // M2CM10 Alarm
        [33].7   // M2CM07 Faulted
        [41]   // M2CM09 Drive Status
        [37].3   // M2CM08 Actual Direction
        [38]   // M2CM08 Speed Reference
        [35]   // M2CM07 A1 Data Out
        [35].1   // M2CM07 Reference ID
        [36]   // M2CM07 A2 Data Out
        [41].8   // M2CM09 At Speed
        [37].0   // M2CM08 Enabled
        [37].1   // M2CM08 Running
        [41].11   // M2CM09 Local Adaptor ID
        [45].10   // M2CM10 Local Adaptor ID
        [37].13   // M2CM08 Reference ID
        [37].14   // M2CM08 Reference ID
        [37].15   // M2CM08 Reference ID
        [41].12   // M2CM09 Reference ID
        [41].2   // M2CM09 Cmd Direction
        [37].9   // M2CM08 Local Adaptor ID
        [37].4   // M2CM08 Accelerating
        [37].5   // M2CM08 Decelerating
        [49].6   // M2CM11 Alarm
        [37].7   // M2CM08 Faulted
        [45]   // M2CM10 Drive Status
        [41].3   // M2CM09 Actual Direction
        [42]   // M2CM09 Speed Reference
        [39]   // M2CM08 A1 Data Out
        [39].5   // M2CM08 Reference ID
        [40]   // M2CM08 A2 Data Out
        [45].8   // M2CM10 At Speed
        [41].0   // M2CM09 Enabled
        [41].1   // M2CM09 Running
        [45].11   // M2CM10 Local Adaptor ID
        [49].10   // M2CM11 Local Adaptor ID
        [41].13   // M2CM09 Reference ID
        [41].14   // M2CM09 Reference ID
        [41].15   // M2CM09 Reference ID
        [45].12   // M2CM10 Reference ID
        [45].2   // M2CM10 Cmd Direction
        [41].9   // M2CM09 Local Adaptor ID
        [41].4   // M2CM09 Accelerating
        [41].5   // M2CM09 Decelerating
        [53].6   // M2CM12 Alarm
        [41].7   // M2CM09 Faulted
        [49]   // M2CM11 Drive Status
        [45].3   // M2CM10 Actual Direction
        [46]   // M2CM10 Speed Reference
        [43]   // M2CM09 A1 Data Out
        [43].9   // M2CM09 Reference ID
        [44]   // M2CM09 A2 Data Out
        [49].8   // M2CM11 At Speed
        [45].0   // M2CM10 Enabled
        [45].1   // M2CM10 Running
        [49].11   // M2CM11 Local Adaptor ID
        [53].10   // M2CM12 Local Adaptor ID
        [45].13   // M2CM10 Reference ID
        [45].14   // M2CM10 Reference ID
        [45].15   // M2CM10 Reference ID
        [47].13   // M2CM10 Reference ID
        [49].2   // M2CM11 Cmd Direction
        [45].9   // M2CM10 Local Adaptor ID
        [45].4   // M2CM10 Accelerating
        [45].5   // M2CM10 Decelerating
        [9].0   // M2CM01 Enabled
        [45].7   // M2CM10 Faulted
        [53]   // M2CM12 Drive Status
        [49].3   // M2CM11 Actual Direction
        [50]   // M2CM11 Speed Reference
        [47]   // M2CM10 A1 Data Out
        [49].12   // M2CM11 Reference ID
        [48]   // M2CM10 A2 Data Out
        [53].8   // M2CM12 At Speed
        [49].0   // M2CM11 Enabled
        [49].1   // M2CM11 Running
        [53].11   // M2CM12 Local Adaptor ID
        [49].13   // M2CM11 Reference ID
        [49].14   // M2CM11 Reference ID
        [49].15   // M2CM11 Reference ID
        [53].12   // M2CM12 Reference ID
        [53].2   // M2CM12 Cmd Direction
        [49].9   // M2CM11 Local Adaptor ID
        [49].4   // M2CM11 Accelerating
        [49].5   // M2CM11 Decelerating
        [9].1   // M2CM01 Running
        [49].7   // M2CM11 Faulted
        [53].3   // M2CM12 Actual Direction
        [54]   // M2CM12 Speed Reference
        [51]   // M2CM11 A1 Data Out
        [52]   // M2CM11 A2 Data Out
        [52].1   // M2CM11 Reference ID
        [53].0   // M2CM12 Enabled
        [53].1   // M2CM12 Running
        [53].13   // M2CM12 Reference ID
        [53].14   // M2CM12 Reference ID
        [53].15   // M2CM12 Reference ID
        [9].3   // M2CM01 Actual Direction
        [53].9   // M2CM12 Local Adaptor ID
        [53].4   // M2CM12 Accelerating
        [53].5   // M2CM12 Decelerating
        [9].7   // M2CM01 Faulted
        [53].7   // M2CM12 Faulted
        [9].10   // M2CM01 Local Adaptor ID
        [9].2   // M2CM01 Cmd Direction
        [55]   // M2CM12 A1 Data Out
        [56]   // M2CM12 A2 Data Out
        [56].5   // M2CM12 Reference ID
        [7]   // RIO SN READ DATA Reserved Fault Table
        [8]   // RIO SN READ DATA Reserved Fault Table
        [9]   // M2CM01 Drive Status
        [9].11   // M2CM01 Local Adaptor ID
        [9].12   // M2CM01 Reference ID
        [9].13   // M2CM01 Reference ID
        [9].14   // M2CM01 Reference ID
        [9].15   // M2CM01 Reference ID
        [9].9   // M2CM01 Local Adaptor ID
        [9].6   // M2CM01 Alarm
        [9].8   // M2CM01 At Speed
   N95 : DINT[95] := ([4] := 74, [10] := 233, [14] := 60, [18] := 5, [19] := 90, [23] := 484, [30] := 200, [31] := 40, [32] := 465, [35] := 212, [36] := 212, [37] := 470, [38] := 465, [40] := 316, [42] := 158, [43] := 228, [44] := 18, [90] := 465, [91] := 470);
        [30]   // PEG SAMPLE Line Speed for Positioning Calculation [(in/sec) * 10]
        [21]   // Stress Sample Transfer Control State Machine
        [43]   // 400 DECK Leadedge Positioning Counter Target
        [38]   // PEG SAMPLE TE Stopping Setpoint for Glass = 60 In [inches x 10]
        [40]   // 400 DECK Dist to Centerline of Stopped Cap from Reliance Handoff eye [in]
        [4].4   // One Shot
        [5].1   // 400 Deck Plate entry in Progress Operate drives At trim speed
        [4].5   // One Shot
        [4].6   // One Shot
        [5].3   // 400 Deck
        [5].4   // 400 Deck
        [5].5   // 400 Deck
        [5].6   // 400 Deck
        [5].7   // 400 Deck
        [6].1   // 400 Deck Conveyor 1 Operate at Trim speed
        [6].2   // 400 Deck Conveyor 2 Operate at Trim speed
        [6].3   // 400 Deck Conveyor 3 Operate at Trim speed
        [6].4   // 400 Deck Conveyor 4 Operate at Trim speed
        [6].5   // 400 Deck Conveyor 5 Operate at Trim speed
        [6].6   // 400 Deck Conveyor 6 Operate at Trim speed
        [6].7   // 400 Deck Conveyor 7 Operate at Trim speed
        [6].8   // 400 Deck Conveyor 8 Operate at Trim speed
        [36]   // PEG SAMPLE TIME ELAPSED FOR CURRENT SAMPLE POSITIONING
        [91]   // PEG SAMPLE Trailedge (HI SPD) Stopping Setpoint [inches x 10]
        [12]   // Sapmle/Peg CAP ID Storage Register
        [5].0   // 400 Deck Plate entry In progress
        [5].2   // 400 Deck Movement in Progress Do not operate Drives
        [44]   // 400 DECK OP Adjust Distance For Larger Plates [in]
